FUNCTION_BLOCK "SINAMICS_LinearPos_ControlTorque"   // FB58, LAD
TITLE = Sinamics drive manager
{ S7_Optimized_Access := 'FALSE' }
AUTHOR : Armitano
VERSION : 1.5
// Return value:
// * 0: OK
// Blocking message:
// * group 1 to 9: general error
// * group 10 to 19: system data error
//   * 10: Sinamics input/output addresses wrong or not setted
//   * 11: Maximum speed in Rpm wrong or not setted
//   * 12: Conversion coefficent for Rpm/mmMin wrong or not setted
//   * 13: Conversion coefficent for mmMin/Rpm wrong or not setted
//   * 14: Maximum acceleration wrong or not setted
//   * 15: Maximum deceleration wrong or not setted
//   * 19: Comunication telegram number unknown
// Warning message:
// * group 20 to 29: user data error
//   * 20: Reference cam signal + reference zero signal no possible
//   * 21: Run command + reverse command no possible
//   * 22: Preset speed at zero during run/reverse command
//   * 23: Run/reverse command during homing command no possible
//   * 24: Absolute positioining no possible without axes referenced
//   * 25: Preset override at zero during run/reverse command
// Other:
// * group 30 to 32: preset data error
//   * 30: Error during send preset value (Check parameters in Sys_Data)
//   * 31: Error during preset command (Check parameters in Sys_Data)
//   * 32: Error during saving preset command (Check Sys_Data)
//   * 34: Error during send preset homing (Check parameters in Sys_Data)
//   * 40: Error during request misured values (Check Sys_Data)
//   * 41: Error during response misured values (Check Sys_Data)
// * group 8000 to 9000: SFC20 code (Read the SFC20 Help)
   VAR_INPUT
      IN_xDrive_EN : Bool;   // Drive enable
      IN_xRun : Bool;   // Run forward
      IN_xReverse : Bool;   // Run backward
      IN_xPositioning : Bool;   // Positioning enable
      IN_xResetFaults : Bool;   // Reset faults
      IN_dSpeed_mm_min : DInt;   // Speed reference [mm/min]
   END_VAR
   VAR_OUTPUT
      OUT_xFeedback : Bool;   // Feedback active
      OUT_xFaultPresent : Bool;   // Fault present
      OUT_iFaultCode : Int;   // Fault code
      OUT_iRetVal : Int;   // Return value in case of wrong configuration
   END_VAR
   VAR
      STC_tUSER_DATA : Struct   // User data (Extended functions commands for execute the application desired)
         tR : Struct
            xReadyfForSwitchOn : Bool;   // Ready for switch on
            xReadyToMove : Bool;   // Ready to move
            xAxleRefered : Bool;   // Axle referenced (only positioner)
            xPositionReached : Bool;   // Position reached (only positioner)
            xAlarmPresent : Bool;   // Alarm present
            xAxleToZero : Bool;   // Axle to zero value (only positioner)
            xAxleAcc : Bool;   // Axle in acceleration
            xAxleDec : Bool;   // Axle in deceleration
            iAlarmCode : Int;   // Alarm code
            dActualPosition_dmm : DInt;   // Actual position value [mm/10] (only positioner)
            dActualSpeed_mm_min : DInt;   // Actual speed value [mm/min]
         END_STRUCT;
         tW : Struct
            xSafetyStop : Bool;   // Safety stop (OFF3)
            xFlyChange : Bool;   // Fly change (only positioner)
            xPH_Select : Bool;   // Photocell selection (only positioner)
            xStartCountOnHead : Bool;   // Start count on glass head (only positioner)
            xStartCountOnTail : Bool;   // Start count on glass tail (only positioner)
            xBrakeRelease : Bool;   // Brake release
            xResetCount : Bool;   // Reset counter (only positioner)
            xPresetRq : Bool;   // Preset request (only absolute encoder)
            xHomeSearch : Bool;   // Home search cycle (only for homing)
            xReverseHoming : Bool;   // Reverse homing search direction (only for homing)
            xReferenceCam : Bool;   // Sensor reference cam for homing cycle + zero mark (only for homing)
            xReferenceZero : Bool;   // Sensor reference zero for homing cycle (only for homing)
            xMDI_Continue : Bool;   // MDI movement continue (only for gearing axes)
            x14 : Bool;
            xHwLimitsEnable : Bool;   // Hardware limits activation (only positioner)
            xEdgePulseStartCount : Bool;   // Edge pulse of start count photocell (for positioning with photocell)
            iOverride_perc : Int := 100;   // Override [%] (only positioner)
            dTarget_dmm : DInt;   // Target position [mm/10] (only positioner)
            dPreset_dmm : DInt;   // Preset position [mm/10] (only for homing & absolute encoder)
            rAcc : Real;   // Acceleration [Pos=m/s2,OpLoop=s]
            rDec : Real;   // Deceleration [Pos=m/s2,OpLoop=s]
         END_STRUCT;
      END_STRUCT;
      STC_tSYS_DATA : Struct   // System data (Info about applications type and HW config.)
         iIOAddress_MM : Int := -1;   // Input/Output addresses for motor module
         iPZD_MM : Int;   // Type of telegram in motor module [111=Positioner, 1=Open/close loop]
         i3 : Int;
         iDiagAddress : Int;   // Diagnostic address of SINAMICS module (only for absolute encoder & homing)
         iPosPZD_CU : Int;   // Number of PZD position in SINAMICS configuration [1,2,3..] (for absolute enc.)
         iPosPZD_MM : Int;   // Number of PZD position in SINAMICS configuration [1,2,3..] (for homing & enc.)
         iEncNumb : Int;   // Encoder number for preset position [0=Encoder1,1=Encoder2] (for absolute enc.)
         dMaxSpeed_rpm : DInt;   // MaxSpeed [rpm]
         d9 : DInt;
         dPosWindow_dmm : DInt := L#1;   // Positioning window [mm/10] (only positioner)
         dTorque : DInt;   // Limit torque value [0-100%]
         dSpeed_reference : DInt;   // Speed refence [rpm]
         d13 : DInt;
         rK_rpm_mmMin : Real;   // K Conversion from rpm to mm/min
         rK_mmMin_Rpm : Real;   // K Conversion from mm/min to rpm (only for Open/close loop)
         rMaxAcc : Real;   // MaxAcc [Pos=m/s2,OpClLoop=s]
         rMaxDec : Real;   // MaxDec [Pos=m/s2,OpClLoop=s]
         r18 : Real;
         r19 : Real;
      END_STRUCT;
      STC_tEXT_DATA : Struct   // Extended data (Functions commands for DCC applications)
         tR : Struct
            x0 : Bool;
            x1 : Bool;
            x2 : Bool;
            x3 : Bool;
            x4 : Bool;
            x5 : Bool;
            x6 : Bool;
            x7 : Bool;
            xMisureDone : Bool;   // Misure executed (Only positioner)
            x9 : Bool;
            x10 : Bool;
            x11 : Bool;
            x12 : Bool;
            x13 : Bool;
            x14 : Bool;
            x15 : Bool;
            tMisureVal : Struct   // Misured values with probe
               tRising : Struct   // Positive edge record valueas
                  dP_Edge1_dmm : DInt;   // Rising edge positive misured value 1 [mm/10] (Only positioner)
                  dP_Edge2_dmm : DInt;   // Rising edge positive misured value 2 [mm/10] (Only positioner)
                  dP_Edge3_dmm : DInt;   // Rising edge positive misured value 3 [mm/10] (Only positioner)
                  dP_Edge4_dmm : DInt;   // Rising edge positive misured value 4 [mm/10] (Only positioner)
                  dP_Edge5_dmm : DInt;   // Rising edge positive misured value 5 [mm/10] (Only positioner)
                  dP_Edge6_dmm : DInt;   // Rising edge positive misured value 6 [mm/10] (Only positioner)
               END_STRUCT;
               tFalling : Struct   // Negative edge record valueas
                  dN_Edge1_dmm : DInt;   // Rising edge negative misured value 1 [mm/10] (Only positioner)
                  dN_Edge2_dmm : DInt;   // Rising edge negative misured value 2 [mm/10] (Only positioner)
                  dN_Edge3_dmm : DInt;   // Rising edge negative misured value 3 [mm/10] (Only positioner)
                  dN_Edge4_dmm : DInt;   // Rising edge negative misured value 4 [mm/10] (Only positioner)
                  dN_Edge5_dmm : DInt;   // Rising edge negative misured value 5 [mm/10] (Only positioner)
                  dN_Edge6_dmm : DInt;   // Rising edge negative misured value 6 [mm/10] (Only positioner)
               END_STRUCT;
            END_STRUCT;
            rgdSpare : Array[0..5] of DInt;
         END_STRUCT;
         tW : Struct
            xGearingCtrl : Bool;   // Active gearing mode
            xControlTorque : Bool;   // Active control torque
            x2 : Bool;
            x3 : Bool;
            x4 : Bool;
            xModuleCorrect : Bool;   // Enable module correction (only positioner with turnover endless)
            x6 : Bool;
            x7 : Bool;
            xEnMisProbe : Bool;   // Enable misure probe (Only positioner)
            xRqMisVal : Bool;   // Request misured values (Only positioner)
            x10 : Bool;
            x11 : Bool;
            x12 : Bool;
            x13 : Bool;
            x14 : Bool;
            x15 : Bool;
            d0 : DInt;
            d1 : DInt;
            d2 : DInt;
            d3 : DInt;
            d4 : DInt;
            d5 : DInt;
            d6 : DInt;
            d7 : DInt;
            d8 : DInt;
            d9 : DInt;
            d10 : DInt;
            d11 : DInt;
            rgdSpare : Array[0..5] of DInt;
         END_STRUCT;
      END_STRUCT;
      STC_tST : Struct
         x0 : Bool;   // Positioning Absolute
         x1 : Bool;   // Positioning with photocell
         x2 : Bool;
         x3 : Bool;
         x4 : Bool;
         x5 : Bool;
         x6 : Bool;   // Target = Feedback target
         x7 : Bool;   // Validation position reached with module correction
         x8 : Bool;   // Preset phases in progress
         x9 : Bool;
         x10 : Bool;
         x11 : Bool;   // Axle resetted
         x12 : Bool;
         x13 : Bool;
         x14 : Bool;
         x15 : Bool;
      END_STRUCT;
      STC_tOS_PN : Struct
         x0 : Bool;   // Run
         x1 : Bool;   // Reverse
         x2 : Bool;   // Positioning
         x3 : Bool;   // Fly change
         x4 : Bool;
         x5 : Bool;
         x6 : Bool;   // Waiting photocell signal
         x7 : Bool;   // Position reached
         x8 : Bool;   // Fly referencing active (Positive edge)
         x9 : Bool;   // Fly referencing active (Negative edge)
         x10 : Bool;   // Preset position
         x11 : Bool;
         x12 : Bool;
         x13 : Bool;   // Request misured values
         x14 : Bool;
         x15 : Bool;
      END_STRUCT;
      STC_tOS : Struct
         x0 : Bool;   // Run
         x1 : Bool;   // Reverse
         x2 : Bool;   // Positioning
         x3 : Bool;   // Fly change
         x4 : Bool;
         x5 : Bool;
         x6 : Bool;   // Waiting photocell signal
         x7 : Bool;
         x8 : Bool;   // Fly referencing active
         x9 : Bool;
         x10 : Bool;
         x11 : Bool;
         x12 : Bool;
         x13 : Bool;
         x14 : Bool;
         x15 : Bool;
      END_STRUCT;
      STC_tPH : Struct
         x0 : Bool;   // Positioning initializing
         x1 : Bool;   // Positioning request
         x2 : Bool;   // Fly change waiting
         x3 : Bool;   // Fly change sending
         x4 : Bool;   // Change command waiting
         x5 : Bool;   // Change command request
         x6 : Bool;   // Wait photocell signal
         x7 : Bool;
         x8 : Bool;   // Send encoder value
         x9 : Bool;   // Send preset command
         x10 : Bool;   // Send saving preset command
         x11 : Bool;   // End preset encoder
         x12 : Bool;
         x13 : Bool;   // Request misured values
         x14 : Bool;   // Waiting response values
         x15 : Bool;   // Misured values recived
      END_STRUCT;
      STC_tPROP : Struct
         i0 : Int;   // Previous cycle [ms]
         i1 : Int;
         i2 : Int;   // Override in sending [%]
         d3 : DInt;   // Speed in sending [mm/min]
         d4 : DInt;   // Target in sending [mm/10]
         r5 : Real;   // Acceleration in sending [m/s2]
         r6 : Real;   // Deceleration in sending [m/s2]
         i7 : Int;
         i8 : Int;
         i9 : Int;
         i10 : Int;
         i11 : Int;   // Override in fly change [%]
         d12 : DInt;   // Speed in fly change [mm/min]
         d13 : DInt;   // Target in fly change [mm/10]
         r14 : Real;   // Acceleration in fly change [m/s2]
         r15 : Real;   // Deceleration in fly change [m/s2]
         i16 : Int;
         i17 : Int;
         i18 : Int;
         i19 : Int;
         i20 : Int;
         tmON_feedback_ms : IEC_TIMER;   // Delay feedback [ms]
      END_STRUCT;
      STC_tR_MngSysReg : Struct   // Managment system register
         tST : Struct
            xRead_Request : Bool;
            xDone : Bool;
            xBusy : Bool;
            xError : Bool;
            xSpare4 : Bool;
            xSpare5 : Bool;
            xSpare6 : Bool;
            xSpare7 : Bool;
            ID : Hw_Io;
            dINDEX : DInt;
            uiLEN : UInt;
            dwSTATUS : DWord;
            uiMLEN : UInt;
         END_STRUCT;
         tDATA : Struct
            tRequestValues : Struct
               wRequest_refere_RequestID : Word := W#16#501;   // (Request_referece=01 Alwais=01 )*(RequestID=01 Read Param)
               wAxis_NoOfParameters : Word := W#16#112;   // (Axis=Num.Object)(NoOfParameters=Num of parameter to Read)
               wAttribute_NoOfElements_1 : Word := W#16#1000;   // (Attribute=10 Alwais=10)(NoOfParameters=Num of subparameter to Read)
               iParameter_number_1 : Int := 21700;   // Parameter_number=Number of the parameter
               wSubindex_1 : Word;   // Subindex
               wAttribute_NoOfElements_2 : Word := W#16#1000;   // (Attribute=10 Alwais=10)(NoOfParameters=Num of subparameter to Read)
               iParameter_number_2 : Int := 21701;   // Parameter_number=Number of the parameter
               wSubindex_2 : Word;   // Subindex
               wAttribute_NoOfElements_3 : Word := W#16#1000;   // (Attribute=10 Alwais=10)(NoOfParameters=Num of subparameter to Read)
               iParameter_number_3 : Int := 21702;   // Parameter_number=Number of the parameter
               wSubindex_3 : Word;   // Subindex
               wAttribute_NoOfElements_4 : Word := W#16#1000;   // (Attribute=10 Alwais=10)(NoOfParameters=Num of subparameter to Read)
               iParameter_number_4 : Int := 21703;   // Parameter_number=Number of the parameter
               wSubindex_4 : Word;   // Subindex
               wAttribute_NoOfElements_5 : Word := W#16#1000;   // (Attribute=10 Alwais=10)(NoOfParameters=Num of subparameter to Read)
               iParameter_number_5 : Int := 21704;   // Parameter_number=Number of the parameter
               wSubindex_5 : Word;   // Subindex
               wAttribute_NoOfElements_6 : Word := W#16#1000;   // (Attribute=10 Alwais=10)(NoOfParameters=Num of subparameter to Read)
               iParameter_number_6 : Int := 21705;   // Parameter_number=Number of the parameter
               wSubindex_6 : Word;   // Subindex
               wAttribute_NoOfElements_7 : Word := W#16#1000;   // (Attribute=10 Alwais=10)(NoOfParameters=Num of subparameter to Read)
               iParameter_number_7 : Int := 21712;   // Parameter_number=Number of the parameter
               wSubindex_7 : Word;   // Subindex
               wAttribute_NoOfElements_8 : Word := W#16#1000;   // (Attribute=10 Alwais=10)(NoOfParameters=Num of subparameter to Read)
               iParameter_number_8 : Int := 21713;   // Parameter_number=Number of the parameter
               wSubindex_8 : Word;   // Subindex
               wAttribute_NoOfElements_9 : Word := W#16#1000;   // (Attribute=10 Alwais=10)(NoOfParameters=Num of subparameter to Read)
               iParameter_number_9 : Int := 21714;   // Parameter_number=Number of the parameter
               wSubindex_9 : Word;   // Subindex
               wAttribute_NoOfElement_10 : Word := W#16#1000;   // (Attribute=10 Alwais=10)(NoOfParameters=Num of subparameter to Read)
               iParameter_number_10 : Int := 21715;   // Parameter_number=Number of the parameter
               wSubindex_10 : Word;   // Subindex
               wAttribute_NoOfElement_11 : Word := W#16#1000;   // (Attribute=10 Alwais=10)(NoOfParameters=Num of subparameter to Read)
               iParameter_number_11 : Int := 21716;   // Parameter_number=Number of the parameter
               wSubindex_11 : Word;   // Subindex
               wAttribute_NoOfElement_12 : Word := W#16#1000;   // (Attribute=10 Alwais=10)(NoOfParameters=Num of subparameter to Read)
               iParameter_number_12 : Int := 21717;   // Parameter_number=Number of the parameter
               wSubindex_12 : Word;   // Subindex
            END_STRUCT;
            tResponseValues : Struct   // Positive edge record valueas
               wRequest_refere_RequestID : Word;   // (Request_referece=01 Alwais=01 )*(RequestID=01 Read Param)
               wAxis_NoOfParameters : Word;   // (Axis=Num.Object)(NoOfParameters=Num of parameter to Read)
               wFormat_N_Values_1 : Word;   // (Format Parametr) (Number of values)
               dRecordValue_1 : DInt;
               wFormat_N_Values_2 : Word;   // (Format Parametr) (Number of values)
               dRecordValue_2 : DInt;
               wFormat_N_Values_3 : Word;   // (Format Parametr) (Number of values)
               dRecordValue_3 : DInt;
               wFormat_N_Values_4 : Word;   // (Format Parametr) (Number of values)
               dRecordValue_4 : DInt;
               wFormat_N_Values_5 : Word;   // (Format Parametr) (Number of values)
               dRecordValue_5 : DInt;
               wFormat_N_Values_6 : Word;   // (Format Parametr) (Number of values)
               dRecordValue_6 : DInt;
               wFormat_N_Values_7 : Word;   // (Format Parametr) (Number of values)
               dRecordValue_7 : DInt;
               wFormat_N_Values_8 : Word;   // (Format Parametr) (Number of values)
               dRecordValue_8 : DInt;
               wFormat_N_Values_9 : Word;   // (Format Parametr) (Number of values)
               dRecordValue_9 : DInt;
               wFormat_N_Values_10 : Word;   // (Format Parametr) (Number of values)
               dRecordValue_10 : DInt;
               wFormat_N_Values_11 : Word;   // (Format Parametr) (Number of values)
               dRecordValue_11 : DInt;
               wFormat_N_Values_12 : Word;   // (Format Parametr) (Number of values)
               dRecordValue_12 : DInt;
            END_STRUCT;
         END_STRUCT;
      END_STRUCT;
      STC_tW_MngSysReg : Struct   // Managment system register
         tST : Struct
            xWrite_Request : Bool;
            xDone : Bool;
            xBusy : Bool;
            xError : Bool;
            xSpare4 : Bool;
            xSpare5 : Bool;
            xSpare6 : Bool;
            xSpare7 : Bool;
            ID : Hw_Io;
            dINDEX : DInt;
            uiLEN : UInt;
            dwSTATUS : DWord;
            iSpare : Int;
         END_STRUCT;
         tDATA : Struct
            wRequest_refere_RequestID : Word := W#16#102;   // (Request_referece=01 Alwais=01 )*(RequestID=02 Change Param)
            wAxis_NoOfParameters : Word := W#16#101;   // (Axis=Num.Object)(NoOfParameters=Num of parameter to change)
            wAttribute_NoOfElements : Word := W#16#1001;   // (Attribute=10 Alwais=10)(NoOfParameters=Num of subparameter to Write)
            iParameter_number : Int := 2599;   // Parameter_number=Number of the parameter
            wSubindex : Word;   // Subindex
            wFormat_NoOfValue : Word := W#16#4301;   // (Format_NoOfValue=Format 42=Word 43=Dword)(Num. of value to transfer)
            dwRegisterValue : DWord := DW#16#1;   // Register value
         END_STRUCT;
      END_STRUCT;
      STC_tReadRecord : RDREC;
      STC_tWriteRecord : WRREC;
      STC_tPZD_Pos : Struct   // Motor module positioner telegram 111
         tR : Struct   // READ
            tZSW1 : Struct   // R2089[0].STATUS WORD 1
               x8 : Bool;   // Tracking error in tolerance
               x9 : Bool;   // Control request
               x10 : Bool;   // Target position reached
               x11 : Bool;   // Reference point set
               x12 : Bool;   // Acknowledgment, traversing block activated
               x13 : Bool;   // In_actl < speed threshold value 3
               x14 : Bool;   // Axis accelerating
               x15 : Bool;   // Axis decelerating
               x0 : Bool;   // Ready for switch on
               x1 : Bool;   // Ready
               x2 : Bool;   // Operation enabled
               x3 : Bool;   // Fault present
               x4 : Bool;   // OFF2
               x5 : Bool;   // OFF3
               x6 : Bool;   // Switching on inhibited active
               x7 : Bool;   // Alarm present
            END_STRUCT;
            tPOS_ZSW1 : Struct   // R2089[3].POSITIONER STATUS WORD 2
               x8 : Bool;   // STOP cam minus active
               x9 : Bool;   // STOP cam plus active
               x10 : Bool;   // Jog active
               x11 : Bool;   // Homing procedure active
               x12 : Bool;   // Flying referencing active
               x13 : Bool;   // Traversing block active
               x14 : Bool;   // Setup active
               x15 : Bool;   // MDI active
               x0 : Bool;   // Active traversing block, bit 0
               x1 : Bool;   // Active traversing block, bit 1
               x2 : Bool;   // Active traversing block, bit 2
               x3 : Bool;   // Active traversing block, bit 3
               x4 : Bool;   // Active traversing block, bit 4
               x5 : Bool;   // Active traversing block, bit 5
               x6 : Bool;   // Reserved
               x7 : Bool;   // Reserved
            END_STRUCT;
            tPOS_ZSW2 : Struct   // R2089[4].POSITIONER STATUS WORD 3
               x8 : Bool;   // Position actual value <= cam switching position 1
               x9 : Bool;   // Position actual value <= cam switching position 2
               x10 : Bool;   // Direct output 1 via traversing block
               x11 : Bool;   // Direct output 2 via traversing block
               x12 : Bool;   // Fixed stop reached
               x13 : Bool;   // Fixed stop clamping torque reached
               x14 : Bool;   // Travel to fixed stop active
               x15 : Bool;   // Traversing command active
               x0 : Bool;   // Tracking mode active
               x1 : Bool;   // Velocity limit active
               x2 : Bool;   // Setpoint available
               x3 : Bool;   // Printing mark outside outer window
               x4 : Bool;   // Axis moves forwards
               x5 : Bool;   // Axis moves backwards
               x6 : Bool;   // Software limit switch minus reached
               x7 : Bool;   // Software limit switch plus reached
            END_STRUCT;
            dFDB_TARGET : DInt;   // R2060[5].Feedback target
            dXIST_A : DInt;   // R2521[0].Actual position value
            dNIST_B : DInt;   // R63.Actual speed value
            iFAULT_CODE : Int;   // R2131.Actual fault code
            iWARN_CODE : Int;   // R2132.Actual alarm code
            iUser : Int;
         END_STRUCT;
         tW : Struct   // WRITE
            tSTW1 : Struct   // CONTROL WORD 1
               x8 : Bool;   // P2589.EPOS jog 1 signal source
               x9 : Bool;   // P2590.EPOS jog 2 signal source
               x10 : Bool;   // P854[0].Control by PLC
               x11 : Bool;   // P2595.EPOS referencing start
               x12 : Bool;   // R2090[12].Enable misure probe
               x13 : Bool;   // P2633.EPOS external block change
               x14 : Bool;   // R2090[14].Gearing_mode
               x15 : Bool;   // P855[0].Brake release
               x0 : Bool;   // P840[0].ON/OFF
               x1 : Bool;   // P844[0].OFF2
               x2 : Bool;   // P848[0].OFF3
               x3 : Bool;   // P852[0].Enable operation
               x4 : Bool;   // P2641.EPOS abort traversing task
               x5 : Bool;   // P2640.EPOS intermediate STOP
               x6 : Bool;   // P2631.EPOS activate traversing task
               x7 : Bool;   // P2103.Acknowledge faults
            END_STRUCT;
            tPOS_STW1 : Struct   // POSITIONER CONTROL WORD 2
               x8 : Bool;   // P2648.EPOS direct setpoint input/MDI positioning type
               x9 : Bool;   // P2651.EPOS direct setpoint input/MDI direction selection positive
               x10 : Bool;   // P2652.EPOS direct setpoint input/MDI direction selection negative
               x11 : Bool;   // P1142[0].Enable reference value
               x12 : Bool;   // P2649.EPOS direct setpoint input/MDI transfer type selection
               x13 : Bool;   // Reserved
               x14 : Bool;   // P2653.EPOS direct setpoint input/MDI setting-up selection
               x15 : Bool;   // P2647.EPOS direct setpoint input/MDI selection
               x0 : Bool;   // P2525.EPOS traversing block selection, bit 0
               x1 : Bool;   // P2526.EPOS traversing block selection, bit 1
               x2 : Bool;   // P2527.EPOS traversing block selection, bit 2
               x3 : Bool;   // P2528.EPOS traversing block selection, bit 3
               x4 : Bool;   // P2529.EPOS traversing block selection, bit 4
               x5 : Bool;   // P2530.EPOS traversing block selection, bit 5
               x6 : Bool;   // P2550.EPOS Enabled control position
               x7 : Bool;   // P2577.EPOS module correction activation
            END_STRUCT;
            tPOS_STW2 : Struct   // POSITIONER CONTROL WORD 3
               x8 : Bool;   // P2597.EPOS referencing type selection
               x9 : Bool;   // P2604.EPOS search for reference, start direction
               x10 : Bool;   // P2510.LR selecting measuring probe evaluation
               x11 : Bool;   // P2511.LR measuring probe evaluation edge
               x12 : Bool;   // Reserved
               x13 : Bool;   // Reserved
               x14 : Bool;   // P2582.EPOS software limit switch activation
               x15 : Bool;   // P2568.EPOS STOP cam activation
               x0 : Bool;   // P2655.EPOS select tracking mode
               x1 : Bool;   // P2596.EPOS set reference point
               x2 : Bool;   // P2612.EPOS search for reference cam
               x3 : Bool;   // Reserved
               x4 : Bool;   // Reserved
               x5 : Bool;   // P2591.EPOS jogging incremental
               x6 : Bool;   // Reserved
               x7 : Bool;   // Reserved
            END_STRUCT;
            iSTW2 : Int;   // P2045.CONTROL WORD 4
            iOVERRIDE : Int;   // P2646.Override % [0-16384]
            dMDI_TARPOS : DInt;   // P2642.Target position for MDI
            dMDI_VELOCITY : DInt;   // P2643.Speed reference for MDI
            iMDI_ACC : Int;   // P2644.Acceleration ramp % for MDI [0-16384]
            iMDI_DEC : Int;   // P2645.Deceleration ramp % for MDI [0-16384]
            iUser : Int;
            iLimitTorque : Int;   // P1528/P1529. Limit torque % [0-16384]
            iReference_Speed : Int;   // P1070. Speed reference % [0-16384]
         END_STRUCT;
      END_STRUCT;
      STC_tPZD_OpCLLoop : Struct   // Motor module open/close loop telegram 1
         tR : Struct   // READ
            tZSW1 : Struct   // R2089[0].STATUS WORD 1
               x8 : Bool;   // Speed setp-act val deviation in tollerance
               x9 : Bool;   // Control request
               x10 : Bool;   // F or n comparision value reached or exceeded
               x11 : Bool;   // Tourque limit reached
               x12 : Bool;   // Open holding brake
               x13 : Bool;   // Alarm motor overtemperature
               x14 : Bool;   // n_act>=0
               x15 : Bool;   // Alarm power unit thermal overload
               x0 : Bool;   // Ready for switch on
               x1 : Bool;   // Ready
               x2 : Bool;   // Operation enabled
               x3 : Bool;   // Fault present
               x4 : Bool;   // OFF2
               x5 : Bool;   // OFF3
               x6 : Bool;   // Switching on inhibited active
               x7 : Bool;   // Alarm present
            END_STRUCT;
            iNIST_A : Int;   // R63.Actual speed value
            iFAULT_CODE : Int;   // R2131.Actual fault code
            iWARN_CODE : Int;   // R2132.Actual alarm code
         END_STRUCT;
         tW : Struct   // WRITE
            tSTW1 : Struct   // CONTROL WORD 1
               x8 : Bool;   // Reserved
               x9 : Bool;   // Reserved
               x10 : Bool;   // P854[0].Control by PLC
               x11 : Bool;   // P1113[0].Setpoint inversion
               x12 : Bool;   // Reserved
               x13 : Bool;   // P1035[0].Motorized potentiometer setpoint raise
               x14 : Bool;   // P1036[0].Motorized potentiometer setpoint lower
               x15 : Bool;   // P855[0] Brake release
               x0 : Bool;   // P840[0].ON/OFF
               x1 : Bool;   // P844[0].OFF2
               x2 : Bool;   // P848[0].OFF3
               x3 : Bool;   // P852[0].Enable operation
               x4 : Bool;   // P1140[0].Enable ramp function generator
               x5 : Bool;   // P1141[0].Continue ramp function generator
               x6 : Bool;   // P1142[0].Enable setpoint
               x7 : Bool;   // P2103[0].Acknowledge faults
            END_STRUCT;
            iNSOLL_A : Int;   // P1070[0].Main set point
            iACC : Int;   // P1138[0].Acceleration ramp % [0-16384]
            iDEC : Int;   // P1139[0].Deceleration ramp % [0-16384]
            iTorque : Int;   // P1528[0].LimitTorqueSuoerior
         END_STRUCT;
      END_STRUCT;
   END_VAR
   VAR_TEMP
      TMP_dOldValue_AR1 : DInt;
      TMP_dOldValue_AR2 : DInt;
      TMP_x : Bool;
      TMP_i : Int;
      TMP_d : DInt;
      TMP_r : Real;
      TMP_a : ANY;
      TMP_dZero : DInt;
      TMP_xAlwaysON : Bool;
      TMP_rActualSpeed : Real;
      TMP_iAddressLength : Int;
      TMP_dActualPosMin_dmm : DInt;   // Actual position minimum tollerance [mm/10]
      TMP_dActualPosMax_dmm : DInt;   // Actual position maximum tollerance [mm/10]
      TMP_iRetVal : Int;
   END_VAR
   VAR_TEMP   // added for the SCL form of the ladder/FBD networks
      _w1 : Bool;
      _w2 : Bool;
      _w3 : Bool;
      _w4 : Bool;
      _w5 : Bool;
      _w6 : Bool;
      _w7 : Bool;
      _w8 : Bool;
      _w9 : Bool;
      _w10 : Bool;
      _w11 : Bool;
      _w12 : Bool;
      _w13 : Bool;
   END_VAR
BEGIN

REGION Network 1 (STL): Save AR1 & AR2 value
   //    TAR1
   //    T     #TMP_dOldValue_AR1
   //    TAR2
   //    T     #TMP_dOldValue_AR2
END_REGION

REGION Network 2: #####_COSTANTS_#####
END_REGION

REGION Network 3 (STL): Initializing
         SET;
         S     #TMP_xAlwaysON;

         L     DINT#0;
         T     #TMP_dZero;

         CALL  FILL
         ( BVAL    := #TMP_dZero,
           RET_VAL := #TMP_iRetVal,
           BLK     := #STC_tPZD_Pos.tR
         );

         CALL  FILL
         ( BVAL    := #TMP_dZero,
           RET_VAL := #TMP_iRetVal,
           BLK     := #STC_tPZD_OpCLLoop.tR
         );

         CALL  FILL
         ( BVAL    := #TMP_dZero,
           RET_VAL := #TMP_iRetVal,
           BLK     := #STC_tW_MngSysReg
         );

         CALL  FILL
         ( BVAL    := #TMP_dZero,
           RET_VAL := #TMP_iRetVal,
           BLK     := #STC_tR_MngSysReg.tST
         );
END_REGION

REGION Network 4: #####_MOTOR_MODULE_#####
END_REGION

REGION Network 5 (STL): Check system data coerence
         L     #STC_tSYS_DATA.iIOAddress_MM;
         L     0;
         <I;
         L     10;
         JC    Err;

         L     #STC_tSYS_DATA.dMaxSpeed_rpm;
         L     DINT#0;
         <=D;
         L     11;
         JC    Err;

         L     #STC_tSYS_DATA.rK_rpm_mmMin;
         L     0.0;
         <=R;
         L     12;
         JC    Err;

         L     #STC_tSYS_DATA.iPZD_MM;
         L     1;
         ==I;
         A(;
         L     #STC_tSYS_DATA.rK_mmMin_Rpm;
         L     0.0;
         <=R;
         );
         L     13;
         JC    Err;

         L     #STC_tSYS_DATA.rMaxAcc;
         L     0.0;
         <=R;
         L     14;
         JC    Err;

         L     #STC_tSYS_DATA.rMaxDec;
         L     0.0;
         <=R;
         L     15;
         JC    Err;

         L     #STC_tSYS_DATA.iPZD_MM;
         L     111;
         ==I;
         L     12;
         T     #TMP_iAddressLength;
         JC    RIn;
         L     #STC_tSYS_DATA.iPZD_MM;
         L     1;
         ==I;
         L     4;
         T     #TMP_iAddressLength;
         JC    RIn;

         L     19;
         JU    Err;

   RIn:  NOP   0;

   //Compute destination position
         L;
         LAR1;
   //byte 1 = 10h (FIXED for S7)
         L     B#16#10;
         T     B[AR1, P#0.0];
   //byte 2 = data type
         L     B#16#4;  //4 = word
         T     B[AR1, P#1.0];
   //byte 3 & 4 = number of element
         L     #TMP_iAddressLength;  //Production data
         T     W[AR1, P#2.0];
   //byte 5 & 6 = number of DB
         L     0;  //DB production data
         T     W[AR1, P#4.0];
   //byte 7 = memory area
         L     B#16#81;  //81h = I (Input)
         T     B[AR1, P#6.0];
   //byte 8 & 9 = address. Bit 0,1,2 of tenth byte is bit offset
   //byte 7 = address (high). Valid value = 0-7. Bit 3,4,5,6,7 always 0

         L     #STC_tSYS_DATA.iIOAddress_MM;  //Item size
         SLW   3;
         T     W[AR1, P#8.0];
         SRD   16;
         AW    16#0007;
         T     B[AR1, P#7.0];

         L     #STC_tSYS_DATA.iPZD_MM;
         L     111;
         ==I;
         JC    T111;

         L     #STC_tSYS_DATA.iPZD_MM;
         L     1;
         ==I;
         JC    T1;

         BEU;
END_REGION

REGION Network 6: #########################_POSITIONER_###########################
END_REGION

REGION Network 7: #####_MATCH_#####
END_REGION

REGION Network 8 (STL): Input copy
   T111: CALL  BLKMOV
         ( SRCBLK  := #TMP_a,
           RET_VAL := #TMP_iRetVal,
           DSTBLK  := #STC_tPZD_Pos.tR
         );
END_REGION

REGION Network 9: Status signals
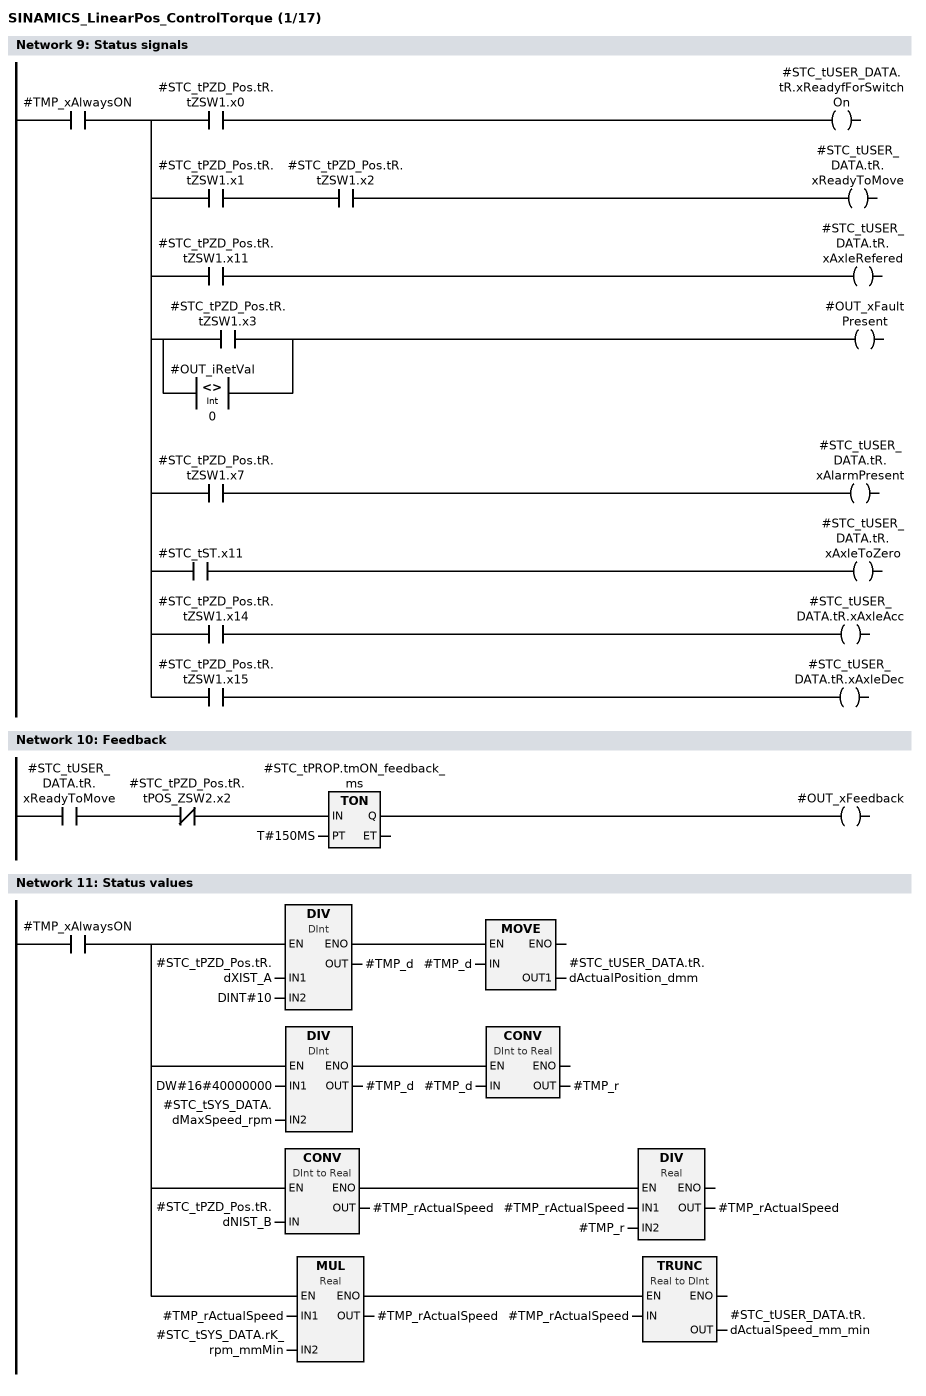
   RUNG wire#powerrail
      Contact( #TMP_xAlwaysON )
      wire#w1
      Contact( #STC_tPZD_Pos.tR.tZSW1.x0 )
      Coil( #STC_tUSER_DATA.tR.xReadyfForSwitchOn )
   END_RUNG
   RUNG wire#w1
      Contact( #STC_tPZD_Pos.tR.tZSW1.x1 )
      Contact( #STC_tPZD_Pos.tR.tZSW1.x2 )
      Coil( #STC_tUSER_DATA.tR.xReadyToMove )
   END_RUNG
   RUNG wire#w1
      Contact( #STC_tPZD_Pos.tR.tZSW1.x11 )
      Coil( #STC_tUSER_DATA.tR.xAxleRefered )
   END_RUNG
   RUNG wire#w1
      Contact( #STC_tPZD_Pos.tR.tZSW1.x3 )
      wire#w2
      Coil( #OUT_xFaultPresent )
   END_RUNG
   RUNG wire#w1
      { S7_Templates := "SrcType := Int" } NE_Contact(in1 := #OUT_iRetVal, in2 := 0)
   END_RUNG wire#w2
   RUNG wire#w1
      Contact( #STC_tPZD_Pos.tR.tZSW1.x7 )
      Coil( #STC_tUSER_DATA.tR.xAlarmPresent )
   END_RUNG
   RUNG wire#w1
      Contact( #STC_tST.x11 )
      Coil( #STC_tUSER_DATA.tR.xAxleToZero )
   END_RUNG
   RUNG wire#w1
      Contact( #STC_tPZD_Pos.tR.tZSW1.x14 )
      Coil( #STC_tUSER_DATA.tR.xAxleAcc )
   END_RUNG
   RUNG wire#w1
      Contact( #STC_tPZD_Pos.tR.tZSW1.x15 )
      Coil( #STC_tUSER_DATA.tR.xAxleDec )
   END_RUNG
   // the same network as SCL:
   #STC_tUSER_DATA.tR.xReadyfForSwitchOn := #TMP_xAlwaysON AND #STC_tPZD_Pos.tR.tZSW1.x0;
   #STC_tUSER_DATA.tR.xReadyToMove := #TMP_xAlwaysON AND #STC_tPZD_Pos.tR.tZSW1.x1 AND #STC_tPZD_Pos.tR.tZSW1.x2;
   #STC_tUSER_DATA.tR.xAxleRefered := #TMP_xAlwaysON AND #STC_tPZD_Pos.tR.tZSW1.x11;
   #OUT_xFaultPresent := #TMP_xAlwaysON AND (#STC_tPZD_Pos.tR.tZSW1.x3 OR (#OUT_iRetVal <> 0));
   #STC_tUSER_DATA.tR.xAlarmPresent := #TMP_xAlwaysON AND #STC_tPZD_Pos.tR.tZSW1.x7;
   #STC_tUSER_DATA.tR.xAxleToZero := #TMP_xAlwaysON AND #STC_tST.x11;
   #STC_tUSER_DATA.tR.xAxleAcc := #TMP_xAlwaysON AND #STC_tPZD_Pos.tR.tZSW1.x14;
   #STC_tUSER_DATA.tR.xAxleDec := #TMP_xAlwaysON AND #STC_tPZD_Pos.tR.tZSW1.x15;
END_REGION

REGION Network 10: Feedback
   #STC_tPROP.tmON_feedback_ms.TON(IN := #STC_tUSER_DATA.tR.xReadyToMove AND NOT #STC_tPZD_Pos.tR.tPOS_ZSW2.x2,
                           PT := T#150MS);
   #OUT_xFeedback := #STC_tPROP.tmON_feedback_ms.Q;
END_REGION

REGION Network 11: Status values
   RUNG wire#powerrail
      Contact( #TMP_xAlwaysON )
      wire#w1
      { S7_Templates := "SrcType := DInt"; S7_GenerateENO := "TRUE" } Div(in1 := #STC_tPZD_Pos.tR.dXIST_A, in2 := DINT#10, out => #TMP_d)
      { S7_GenerateENO := "TRUE" } Move(in := #TMP_d, out1 => #STC_tUSER_DATA.tR.dActualPosition_dmm)
   END_RUNG
   RUNG wire#w1
      { S7_Templates := "SrcType := DInt"; S7_GenerateENO := "TRUE" } Div(in1 := DW#16#40000000, in2 := #STC_tSYS_DATA.dMaxSpeed_rpm, out => #TMP_d)
      { S7_Templates := "[SrcType := DInt, DestType := Real]"; S7_GenerateENO := "TRUE" } Convert(in := #TMP_d, out => #TMP_r)
   END_RUNG
   RUNG wire#w1
      { S7_Templates := "[SrcType := DInt, DestType := Real]"; S7_GenerateENO := "TRUE" } Convert(in := #STC_tPZD_Pos.tR.dNIST_B, out => #TMP_rActualSpeed)
      { S7_Templates := "SrcType := Real"; S7_GenerateENO := "TRUE" } Div(in1 := #TMP_rActualSpeed, in2 := #TMP_r, out => #TMP_rActualSpeed)
   END_RUNG
   RUNG wire#w1
      { S7_Templates := "SrcType := Real"; S7_GenerateENO := "TRUE" } Mul(in1 := #TMP_rActualSpeed, in2 := #STC_tSYS_DATA.rK_rpm_mmMin, out => #TMP_rActualSpeed)
      { S7_Templates := "[SrcType := Real, DestType := DInt]"; S7_GenerateENO := "TRUE" } Trunc(in := #TMP_rActualSpeed, out => #STC_tUSER_DATA.tR.dActualSpeed_mm_min)
   END_RUNG
   // the same network as SCL:
   // ENO of a box is taken as its EN; it also drops when the box reports an error
   IF #TMP_xAlwaysON THEN
       #TMP_d := #STC_tPZD_Pos.tR.dXIST_A / DINT#10;
       #STC_tUSER_DATA.tR.dActualPosition_dmm := #TMP_d;
       #TMP_d := DW#16#40000000 / #STC_tSYS_DATA.dMaxSpeed_rpm;
       #TMP_r := DINT_TO_REAL(#TMP_d);
       #TMP_rActualSpeed := DINT_TO_REAL(#STC_tPZD_Pos.tR.dNIST_B);
       #TMP_rActualSpeed := #TMP_rActualSpeed / #TMP_r;
       #TMP_rActualSpeed := #TMP_rActualSpeed * #STC_tSYS_DATA.rK_rpm_mmMin;
       #STC_tUSER_DATA.tR.dActualSpeed_mm_min := TRUNC(#TMP_rActualSpeed);
   END_IF;
END_REGION

REGION Network 12: #####_STATUSES_#####
END_REGION

REGION Network 13: Type of positioning
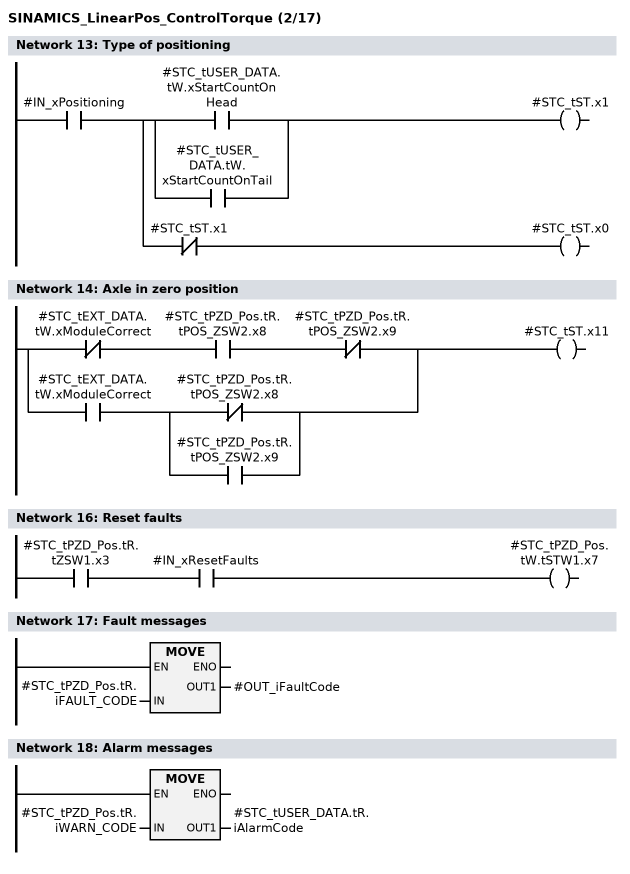
   RUNG wire#powerrail
      Contact( #IN_xPositioning )
      wire#w1
      Contact( #STC_tUSER_DATA.tW.xStartCountOnHead )
      wire#w2
      Coil( #STC_tST.x1 )
   END_RUNG
   RUNG wire#w1
      Contact( #STC_tUSER_DATA.tW.xStartCountOnTail )
   END_RUNG wire#w2
   RUNG wire#w1
      I_Contact( #STC_tST.x1 )
      Coil( #STC_tST.x0 )
   END_RUNG
   // the same network as SCL:
   #STC_tST.x1 := #IN_xPositioning AND (#STC_tUSER_DATA.tW.xStartCountOnHead OR #STC_tUSER_DATA.tW.xStartCountOnTail);
   #STC_tST.x0 := #IN_xPositioning AND NOT #STC_tST.x1;
END_REGION

REGION Network 14: Axle in zero position
   RUNG wire#powerrail
      I_Contact( #STC_tEXT_DATA.tW.xModuleCorrect )
      Contact( #STC_tPZD_Pos.tR.tPOS_ZSW2.x8 )
      I_Contact( #STC_tPZD_Pos.tR.tPOS_ZSW2.x9 )
      wire#w1
      Coil( #STC_tST.x11 )
   END_RUNG
   RUNG wire#powerrail
      Contact( #STC_tEXT_DATA.tW.xModuleCorrect )
      wire#w2
      I_Contact( #STC_tPZD_Pos.tR.tPOS_ZSW2.x8 )
   END_RUNG wire#w1
   RUNG wire#w2
      Contact( #STC_tPZD_Pos.tR.tPOS_ZSW2.x9 )
   END_RUNG wire#w1
   // the same network as SCL:
   #STC_tST.x11 := (NOT #STC_tEXT_DATA.tW.xModuleCorrect AND #STC_tPZD_Pos.tR.tPOS_ZSW2.x8 AND NOT #STC_tPZD_Pos.tR.tPOS_ZSW2.x9) OR (#STC_tEXT_DATA.tW.xModuleCorrect AND (NOT #STC_tPZD_Pos.tR.tPOS_ZSW2.x8 OR #STC_tPZD_Pos.tR.tPOS_ZSW2.x9));
END_REGION

REGION Network 15: #####_ALARMS_#####
END_REGION

REGION Network 16: Reset faults
   RUNG wire#powerrail
      Contact( #STC_tPZD_Pos.tR.tZSW1.x3 )
      Contact( #IN_xResetFaults )
      Coil( #STC_tPZD_Pos.tW.tSTW1.x7 )
   END_RUNG
   // the same network as SCL:
   #STC_tPZD_Pos.tW.tSTW1.x7 := #STC_tPZD_Pos.tR.tZSW1.x3 AND #IN_xResetFaults;
END_REGION

REGION Network 17: Fault messages
   RUNG wire#powerrail
      { S7_GenerateENO := "TRUE" } Move(in := #STC_tPZD_Pos.tR.iFAULT_CODE, out1 => #OUT_iFaultCode)
   END_RUNG
   // the same network as SCL:
   #OUT_iFaultCode := #STC_tPZD_Pos.tR.iFAULT_CODE;
END_REGION

REGION Network 18: Alarm messages
   RUNG wire#powerrail
      { S7_GenerateENO := "TRUE" } Move(in := #STC_tPZD_Pos.tR.iWARN_CODE, out1 => #STC_tUSER_DATA.tR.iAlarmCode)
   END_RUNG
   // the same network as SCL:
   #STC_tUSER_DATA.tR.iAlarmCode := #STC_tPZD_Pos.tR.iWARN_CODE;
END_REGION

REGION Network 19: #####_PHASES_&_LOGICS_#####
END_REGION

REGION Network 20: Enable PLC control